// TIA Portal project "datadiode_receiver" (V17)

(* hardware
DEVICE "S7-1500/ET200MP-Station_1"  S7-1500 station
   slot 0: "Profilschiene_0"  Rack  6ES7 590-1***0-0AA0
   slot 1: "PLC_1"  CPU 1516-3 PN/DP  6ES7 516-3AN02-0AB0  V2.9
      slot 3: "CPU-Display_1"  6ES7591-1BA00-0AA0
      slot 32768: "PROFINET-Schnittstelle_1"  X1
      slot 33024: "PROFINET-Schnittstelle_2"  X2
      slot 33280: "DP-Schnittstelle_1"  X3
      slot 34817: "Virtual CP interface port_1"  Virtual CP interface port  Virtual CP interface port
DEVICE "S7-1500/ET200MP-Station_2"  S7-1500 station
   slot 0: "Profilschiene_0"  Rack  6ES7 590-1***0-0AA0
   slot 1: "workstation5.rio"  IM 155-5 PN ST  6ES7 155-5AA00-0AB0  V3.0
   slot 2: "DI 32x24VDC HF_1"  DI 32x24VDC HF  6ES7 521-1BL00-0AB0  V2.1
   slot 3: "DQ 32x24VDC/0.5A HF_1"  DQ 32x24VDC/0.5A HF  6ES7 522-1BL01-0AB0  V1.0
   slot 4: "AI 8xU/I/RTD/TC ST_1"  AI 8xU/I/RTD/TC ST  6ES7 531-7KF00-0AB0  V2.1
   slot 5: "AQ 8xU/I HS_1"  AQ 8xU/I HS  6ES7 532-5HF00-0AB0  V2.0
DEVICE "GSD-Geraet_1"  GSD.Device.PN
   slot 0: "Baugruppenträger"  Rack  V1.0
   slot 0: "datadiodereceiver"  Datadiodereceiver  123 444 777  V0.1.0
      slot 0: "Datadiodereceiver"  Datadiodereceiver
      slot 1: "X1"  X1
         slot 1: "X1 P1"  X1 P1
      slot 1: "Status module_1"  Status module  1.0
         slot 0: "Status Submodule"  Status Submodule
   slot 2: "Temperature Module_1"  Temperature Module  1.0
      slot 0: "Temperature submodule"  Temperature submodule
   slot 3: "Tank Module_1"  Tank Module  1.0
      slot 0: "tank submodule"  tank submodule
   slot 4: "Flow rate Module_1"  Flow rate Module  1.0
      slot 0: "Flow rate Submodule"  Flow rate Submodule
   slot 5: "Pressure Module_1"  Pressure Module  1.0
      slot 0: "Pressure Submodule"  Pressure Submodule
DEVICE "HMI_1"  KTP700 Basic PN
   slot 0: "HMI_1"  KTP700 Basic PN  6AV2 123-2GB03-0AX0  17.0.0.0
   slot 1: "HMI_RT_1"  KTP700 Basic PN  6AV2 123-2GB03-0AX0  17.0.0.0
   slot 5: "HMI_1.IE_CP_1"  PROFINET Interface  17.0.0.0
      slot 1: "PROFINET Schnittstelle_1"  PROFINET Interface
         slot 1: "Port_1"  Port
*)

// ===== PLC "PLC_1"  CPU 1516-3 PN/DP =====

VAR_GLOBAL   // PLC tag table "Standard-Variablentabelle"
   "StatusLED" AT %Q0.0 : Bool;
   "TemperaturLED" AT %Q0.1 : Bool;
   "TankLED" AT %Q0.2 : Bool;
   "FlowRateLED" AT %Q0.3 : Bool;
   "PressureLED" AT %Q0.4 : Bool;
   "statusVIn" AT %IW20 : UInt;
   "tempVIn" AT %IW22 : UInt;
   "tankVIn" AT %IW24 : UInt;
   "flowrateVIn" AT %ID26 : Real;
   "pressureVIn" AT %ID30 : Real;
END_VAR

DATA_BLOCK "HMICom"   // DB1
{ S7_Optimized_Access := 'TRUE' }
VERSION : 0.1
   VAR
      status : Bool;
      temperatur1 : Bool;
      temperatur2 : Bool;
      temperatur3 : Bool;
      tank1 : Bool;
      tank2 : Bool;
      tank3 : Bool;
      flowrate : Bool;
      pressure : Bool;
   END_VAR
BEGIN
END_DATA_BLOCK

ORGANIZATION_BLOCK "Main"   // OB1, LAD, ProgramCycle
TITLE = "Main Program Sweep (Cycle)"
{ S7_Optimized_Access := 'TRUE' }
VERSION : 0.1
   VAR_INPUT
      Initial_Call : Bool;   // Initial call of this OB
      Remanence : Bool;   // =True, if remanent data are available
   END_VAR
   VAR_TEMP
      status_t : Bool;
      flowrate_t : Bool;
      temperatur_t : Bool;
      tank_t : Bool;
      pressure_t : Bool;
   END_VAR
   VAR CONSTANT
      temp_threshold : UInt := 70;
      tank_threshold : UInt := 100;
      flowrate_threshold : Real := 30.0;
      pressure_threshold : Real := 500.0;
   END_VAR
BEGIN

REGION Network 1 (SCL): needs to be changed look at hardware
   IF "statusVIn" > 0 THEN
       "StatusLED" := TRUE;
       #status_t := TRUE;
   ELSE
       "StatusLED" := FALSE;
       #status_t := FALSE;
   END_IF;
END_REGION

REGION Network 2 (SCL): after you put in the moduls
   IF "tankVIn" > #tank_threshold THEN
       "TankLED" := TRUE;
       #tank_t := TRUE;
   ELSE
       "TankLED" := FALSE;
       #tank_t := FALSE;
   END_IF;
END_REGION

REGION Network 3 (SCL): after you put in the moduls
   IF "flowrateVIn" > #flowrate_threshold THEN
       "FlowRateLED" := TRUE;
       #flowrate_t := TRUE;
   ELSE
       "FlowRateLED" := FALSE;
       #flowrate_t := FALSE;
   END_IF;
END_REGION

REGION Network 4 (SCL): after you put in the moduls
   IF "pressureVIn" > #pressure_threshold THEN
       "PressureLED" := TRUE;
       #pressure_t := TRUE;
   ELSE
       "PressureLED" := FALSE;
       #pressure_t := FALSE;
   END_IF;
END_REGION

REGION Network 5
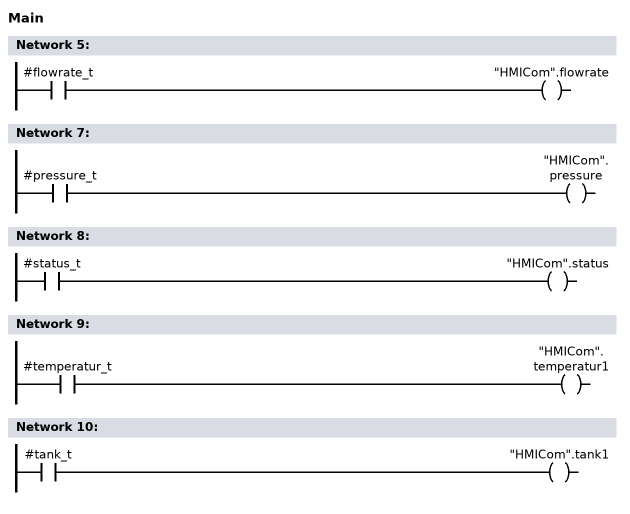
   RUNG wire#powerrail
      Contact( #flowrate_t )
      Coil( "HMICom".flowrate )
   END_RUNG
   // the same network as SCL:
   "HMICom".flowrate := #flowrate_t;
END_REGION

REGION Network 6 (SCL): after you put in the moduls
   IF "tempVIn" > #temp_threshold THEN
       "TemperaturLED" := TRUE;
       #temperatur_t := TRUE;
   ELSE
       "TemperaturLED" := FALSE;
       #temperatur_t := FALSE;
   END_IF;
END_REGION

REGION Network 7
   RUNG wire#powerrail
      Contact( #pressure_t )
      Coil( "HMICom".pressure )
   END_RUNG
   // the same network as SCL:
   "HMICom".pressure := #pressure_t;
END_REGION

REGION Network 8
   RUNG wire#powerrail
      Contact( #status_t )
      Coil( "HMICom".status )
   END_RUNG
   // the same network as SCL:
   "HMICom".status := #status_t;
END_REGION

REGION Network 9
   RUNG wire#powerrail
      Contact( #temperatur_t )
      Coil( "HMICom".temperatur1 )
   END_RUNG
   // the same network as SCL:
   "HMICom".temperatur1 := #temperatur_t;
END_REGION

REGION Network 10
   RUNG wire#powerrail
      Contact( #tank_t )
      Coil( "HMICom".tank1 )
   END_RUNG
   // the same network as SCL:
   "HMICom".tank1 := #tank_t;
END_REGION
END_ORGANIZATION_BLOCK

(* ===== HMI "HMI_RT_1" =====
connection "HMI_Verbindung_1": ETHERNET, SMART_S7_1500_OMS

HMI tags "Standard-Variablentabelle"
   "statusVIn" : UInt = PLC statusVIn AT %IW20, 1 s
   "HMICom_status" : Bool = PLC HMICom.status, 1 s
   "HMICom_tank" : Bool = PLC HMICom.temperatur2, 1 s
   "HMICom_tank1" : Bool = PLC HMICom.tank1, 1 s
   "HMICom_tank2" : Bool = PLC HMICom.tank2, 1 s
   "HMICom_tank3" : Bool = PLC HMICom.tank3, 1 s
   "HMICom_flowrate" : Bool = PLC HMICom.flowrate, 1 s
   "HMICom_pressure" : Bool = PLC HMICom.pressure, 1 s
   "HMICom_temperatur1" : Bool = PLC HMICom.temperatur1, 1 s

screen "Main" 800x480
   Circle "Kreis_1" at 45,35 size 57x57
      Appearance <- "HMICom_status"
   TextField "Textfeld_1" at 116,34 size 104x47; Text 'Status'
   TextField "Textfeld_2" at 610,385 size 71x37; Text 'Tank'
   Circle "Kreis_2" at 45,243 size 57x57
      Appearance <- "HMICom_flowrate"
   Circle "Kreis_3" at 44,318 size 57x57
      Appearance <- "HMICom_pressure"
   TextField "Textfeld_3" at 109,243 size 151x47; Text 'FlowRate'
   TextField "Textfeld_4" at 110,320 size 141x47; Text 'Pressure'
   Rectangle "Rechteck_4" at 539,110 size 206x260
      Appearance <- "HMICom_tank1"
   Circle "Kreis_4" at 42,168 size 57x57
      Appearance <- "HMICom_temperatur1"
   TextField "Textfeld_5" at 116,168 size 210x47; Text 'Temperature'
*)